(* Logix 5000 project; controller PLC_MCC1300_75F1 vendor 1 type 14 code 166 rev 32.11; software revision 32.04; part 19 of 83 *)
(* tags used below, declared in another part *)
   GP_OB_InitializeMain : GP_OB_Initialize;
   M302SpeedUp : MAC_SpeedUp;
   M310_M4_DR_B1 : AXIS_CIP_DRIVE;
   M310_M5_DR_B2 : AXIS_CIP_DRIVE;
   M310B : MAC_Conveyor;
   M310B_Data : UDT_Convoy_SL;
   M310B_M1_DR_IN_MAR : MOTION_INSTRUCTION;
   M310B_M1_DR_IN_MAS : MOTION_INSTRUCTION;
   M310B_M1_DR_OUT_MAJ : MOTION_INSTRUCTION;
   M310B_M1_DR_OUT_MAS : MOTION_INSTRUCTION;
   M310B_M2_DR_IN_MAJ : MOTION_INSTRUCTION;
   M310B_M2_DR_IN_MAR : MOTION_INSTRUCTION;
   M310B_M2_DR_IN_MAS : MOTION_INSTRUCTION;
   M310B_M2_DR_IN_MRP : MOTION_INSTRUCTION;
   M310B_M2_DR_MAFR : MOTION_INSTRUCTION;
   M310B_M2_DR_MDR : MOTION_INSTRUCTION;
   M310B_M2_DR_MSF : MOTION_INSTRUCTION;
   M310B_M2_DR_MSO : MOTION_INSTRUCTION;
   M310B_M2_DR_OUT_MAJ : MOTION_INSTRUCTION;
   M310B_M2_DR_OUT_MAM : MOTION_INSTRUCTION;
   M310B_M2_DR_OUT_MAR : MOTION_INSTRUCTION;
   M310B_M2_DR_OUT_MAS : MOTION_INSTRUCTION;
   M310B_M2_DR_OUT_MCD : MOTION_INSTRUCTION;
   M310B_M2_DR_OUT_MRP : MOTION_INSTRUCTION;
   M310B_SpaceConv_Utilities : SpaceConv_Utilities;
   M310B_xOS_PosReq : BOOL;
   TMP_d : DINT;
   TMP_dDirection : DINT;
   TMP_r : REAL;
   TMP_rAcc : REAL;
   TMP_rDec : REAL;
   TMP_rSpeed : REAL;
   TMP_rTarget_M2 : REAL;
   TMP_xPositioning : BOOL;
   TMP_xPositioning_M2 : BOOL;
   TMP_xReverse : BOOL;
   TMP_xReverse_M1 : BOOL;
   TMP_xReverse_M2 : BOOL;
   TMP_xRun : BOOL;
   TMP_xRun_M1 : BOOL;
   TMP_xRun_M2 : BOOL;
   xAlwaysOFF : BOOL;
   xDebugOFF : BOOL;
   Z300_Conveyor : UDT_StandConv[29];
   Z300_Conveyor_Conf : UDT_Conveyor_Config[29];
   Z300_Conveyor_HMW : MAC_Conveyor_ZC_HMW[29];
   Z300_Conveyor_IN_MOTION : MAC_Conveyor_ZC_IN_MOTION[29];
   Z301_HMR : MAC_Zone_ML_HMR;
   Z401 : MAC_Zone;
(* CommandLogic, continued *)

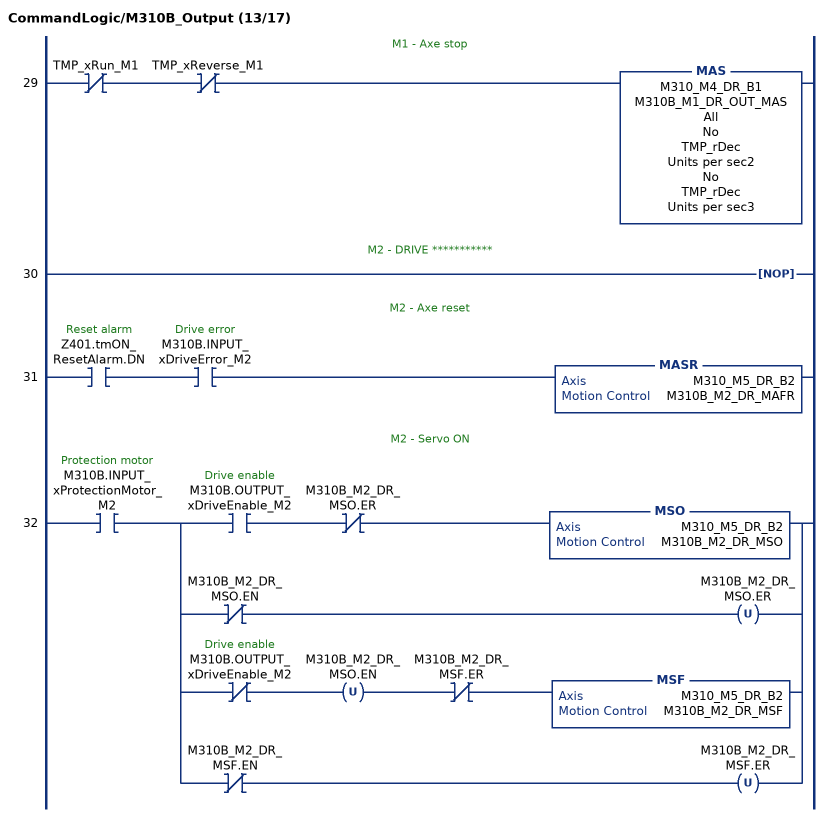
   [picture p150: CommandLogic/M310B_Output rungs 29-32]
   // M1 - Axe stop
   29: XIO(TMP_xRun_M1)XIO(TMP_xReverse_M1)MAS(M310_M4_DR_B1,M310B_M1_DR_OUT_MAS,All,No,TMP_rDec,Units per sec2,No,TMP_rDec,Units per sec3);
   // M2 - DRIVE ***********
   30: NOP();
   // M2 - Axe reset
   31: XIC(Z401.tmON_ResetAlarm.DN)XIC(M310B.INPUT_xDriveError_M2)MASR(M310_M5_DR_B2,M310B_M2_DR_MAFR);
   // M2 - Servo ON
   32: XIC(M310B.INPUT_xProtectionMotor_M2)[XIC(M310B.OUTPUT_xDriveEnable_M2) XIO(M310B_M2_DR_MSO.ER) MSO(M310_M5_DR_B2,M310B_M2_DR_MSO) ,XIO(M310B_M2_DR_MSO.EN) OTU(M310B_M2_DR_MSO.ER) ,XIO(M310B.OUTPUT_xDriveEnable_M2) OTU(M310B_M2_DR_MSO.EN) XIO(M310B_M2_DR_MSF.ER) MSF(M310_M5_DR_B2,M310B_M2_DR_MSF) ,XIO(M310B_M2_DR_MSF.EN) OTU(M310B_M2_DR_MSF.ER) ];
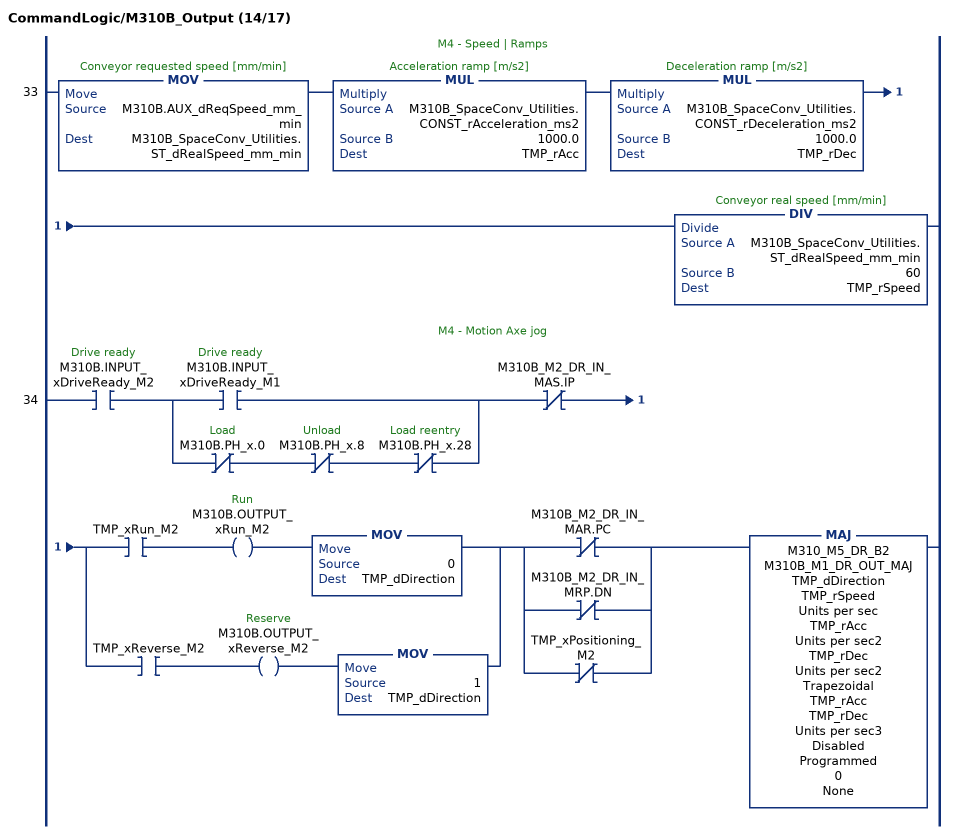
   // M4 - Speed | Ramps
   33: MOV(M310B.AUX_dReqSpeed_mm_min,M310B_SpaceConv_Utilities.ST_dRealSpeed_mm_min)MUL(M310B_SpaceConv_Utilities.CONST_rAcceleration_ms2,1000.0,TMP_rAcc)MUL(M310B_SpaceConv_Utilities.CONST_rDeceleration_ms2,1000.0,TMP_rDec)DIV(M310B_SpaceConv_Utilities.ST_dRealSpeed_mm_min,60,TMP_rSpeed);
   // M4 - Motion Axe jog
   34: XIC(M310B.INPUT_xDriveReady_M2)[XIC(M310B.INPUT_xDriveReady_M1) ,XIO(M310B.PH_x.0) XIO(M310B.PH_x.8) XIO(M310B.PH_x.28) ]XIO(M310B_M2_DR_IN_MAS.IP)[XIC(TMP_xRun_M2) OTE(M310B.OUTPUT_xRun_M2) MOV(0,TMP_dDirection) ,XIC(TMP_xReverse_M2) OTE(M310B.OUTPUT_xReverse_M2) MOV(1,TMP_dDirection) ][XIO(M310B_M2_DR_IN_MAR.PC) ,XIO(M310B_M2_DR_IN_MRP.DN) ,XIO(TMP_xPositioning_M2) ]MAJ(M310_M5_DR_B2,M310B_M1_DR_OUT_MAJ,TMP_dDirection,TMP_rSpeed,Units per sec,TMP_rAcc,Units per sec2,TMP_rDec,Units per sec2,Trapezoidal,TMP_rAcc,TMP_rDec,Units per sec3,Disabled,Programmed,0,None);
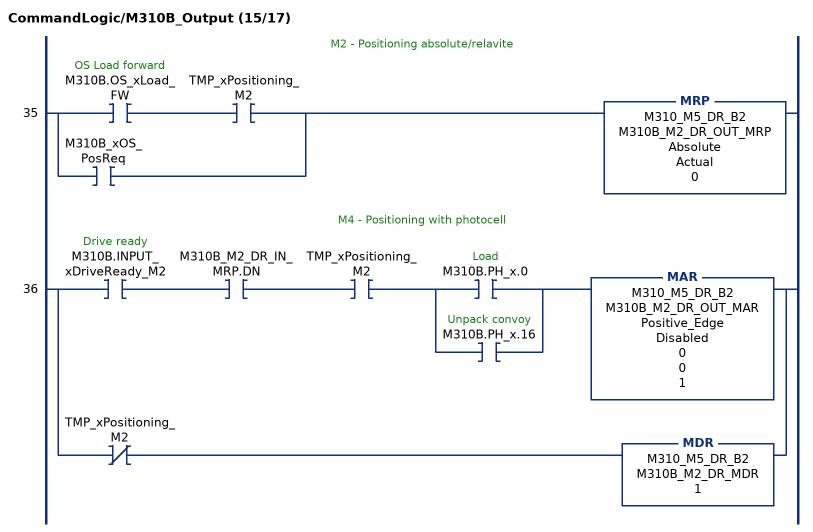
   // M2 - Positioning absolute/relavite
   35: [XIC(M310B.OS_xLoad_FW) XIC(TMP_xPositioning_M2) ,XIC(M310B_xOS_PosReq) ]MRP(M310_M5_DR_B2,M310B_M2_DR_OUT_MRP,Absolute,Actual,0);
   // M4 - Positioning with photocell
   36: [XIC(M310B.INPUT_xDriveReady_M2) XIC(M310B_M2_DR_IN_MRP.DN) XIC(TMP_xPositioning_M2) [XIC(M310B.PH_x.0) ,XIC(M310B.PH_x.16) ] MAR(M310_M5_DR_B2,M310B_M2_DR_OUT_MAR,Positive_Edge,Disabled,0,0,1) ,XIO(TMP_xPositioning_M2) MDR(M310_M5_DR_B2,M310B_M2_DR_MDR,1) ];
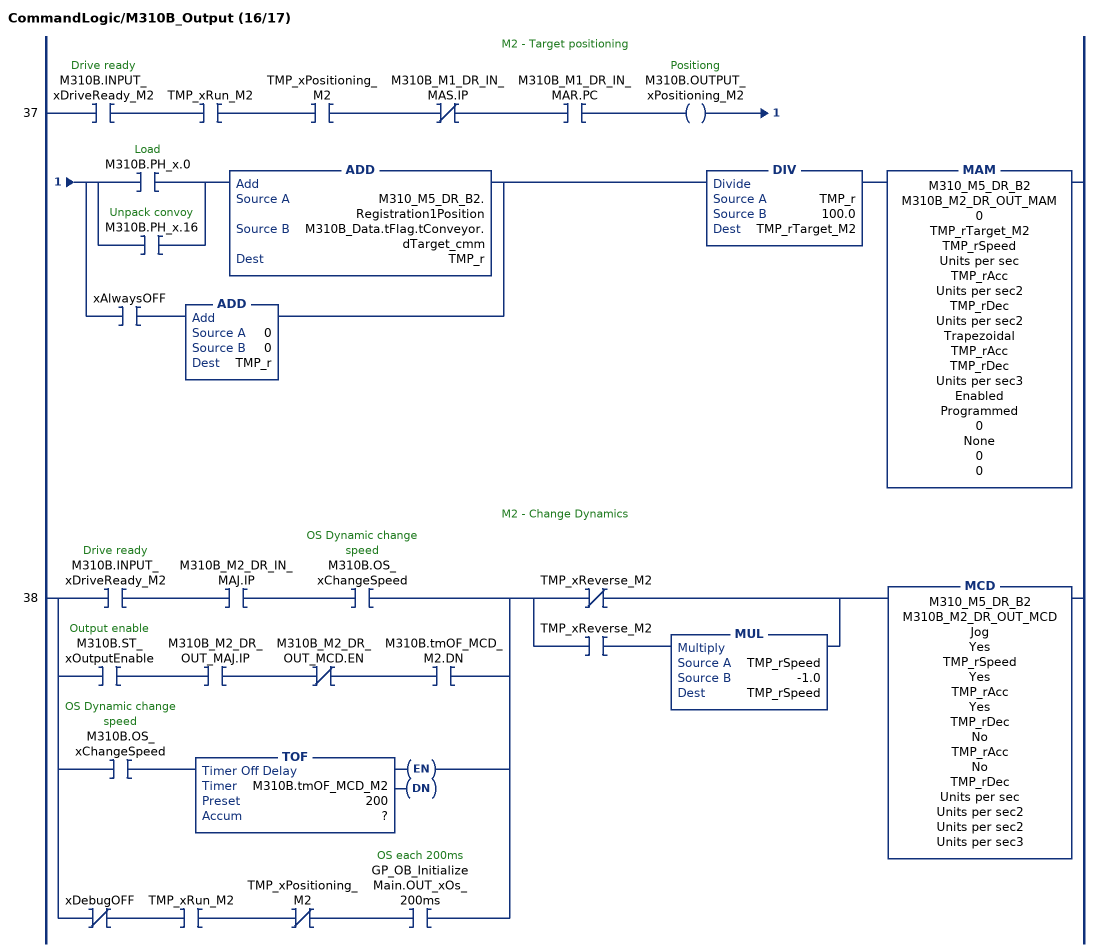
   // M2 - Target positioning
   37: XIC(M310B.INPUT_xDriveReady_M2)XIC(TMP_xRun_M2)XIC(TMP_xPositioning_M2)XIO(M310B_M1_DR_IN_MAS.IP)XIC(M310B_M1_DR_IN_MAR.PC)OTE(M310B.OUTPUT_xPositioning_M2)[[XIC(M310B.PH_x.0) ,XIC(M310B.PH_x.16) ] ADD(M310_M5_DR_B2.Registration1Position,M310B_Data.tFlag.tConveyor.dTarget_cmm,TMP_r) ,XIC(xAlwaysOFF) ADD(0,0,TMP_r) ]DIV(TMP_r,100.0,TMP_rTarget_M2)MAM(M310_M5_DR_B2,M310B_M2_DR_OUT_MAM,0,TMP_rTarget_M2,TMP_rSpeed,Units per sec,TMP_rAcc,Units per sec2,TMP_rDec,Units per sec2,Trapezoidal,TMP_rAcc,TMP_rDec,Units per sec3,Enabled,Programmed,0,None,0,0);
   // M2 - Change Dynamics
   38: [XIC(M310B.INPUT_xDriveReady_M2) XIC(M310B_M2_DR_IN_MAJ.IP) XIC(M310B.OS_xChangeSpeed) ,XIC(M310B.ST_xOutputEnable) XIC(M310B_M2_DR_OUT_MAJ.IP) XIO(M310B_M2_DR_OUT_MCD.EN) XIC(M310B.tmOF_MCD_M2.DN) ,XIC(M310B.OS_xChangeSpeed) TOF(M310B.tmOF_MCD_M2,?,?) ,XIO(xDebugOFF) XIC(TMP_xRun_M2) XIO(TMP_xPositioning_M2) XIC(GP_OB_InitializeMain.OUT_xOs_200ms) ][XIO(TMP_xReverse_M2) ,XIC(TMP_xReverse_M2) MUL(TMP_rSpeed,-1.0,TMP_rSpeed) ]MCD(M310_M5_DR_B2,M310B_M2_DR_OUT_MCD,Jog,Yes,TMP_rSpeed,Yes,TMP_rAcc,Yes,TMP_rDec,No,TMP_rAcc,No,TMP_rDec,Units per sec,Units per sec2,Units per sec2,Units per sec3);
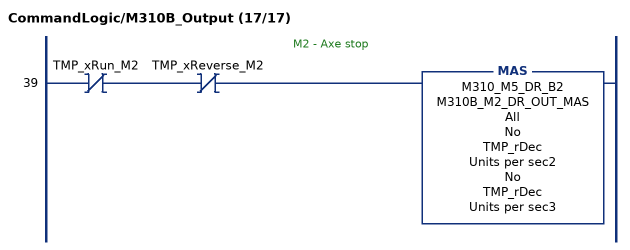
   // M2 - Axe stop
   39: XIO(TMP_xRun_M2)XIO(TMP_xReverse_M2)MAS(M310_M5_DR_B2,M310B_M2_DR_OUT_MAS,All,No,TMP_rDec,Units per sec2,No,TMP_rDec,Units per sec3);
END_ROUTINE

ROUTINE M310M1_Conveyor_Output   (* ladder *)
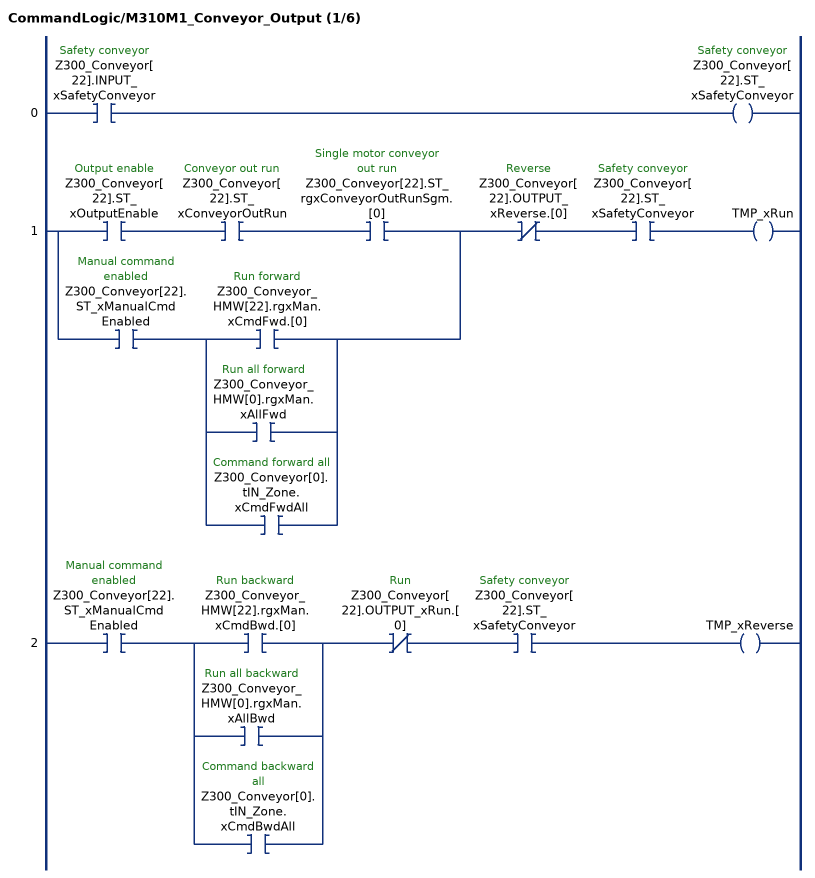
   0: XIC(Z300_Conveyor[22].INPUT_xSafetyConveyor)OTE(Z300_Conveyor[22].ST_xSafetyConveyor);
   1: [XIC(Z300_Conveyor[22].ST_xOutputEnable) XIC(Z300_Conveyor[22].ST_xConveyorOutRun) XIC(Z300_Conveyor[22].ST_rgxConveyorOutRunSgm.[0]) ,XIC(Z300_Conveyor[22].ST_xManualCmdEnabled) [XIC(Z300_Conveyor_HMW[22].rgxMan.xCmdFwd.[0]) ,XIC(Z300_Conveyor_HMW[0].rgxMan.xAllFwd) ,XIC(Z300_Conveyor[0].tIN_Zone.xCmdFwdAll) ] ]XIO(Z300_Conveyor[22].OUTPUT_xReverse.[0])XIC(Z300_Conveyor[22].ST_xSafetyConveyor)OTE(TMP_xRun);
   2: XIC(Z300_Conveyor[22].ST_xManualCmdEnabled)[XIC(Z300_Conveyor_HMW[22].rgxMan.xCmdBwd.[0]) ,XIC(Z300_Conveyor_HMW[0].rgxMan.xAllBwd) ,XIC(Z300_Conveyor[0].tIN_Zone.xCmdBwdAll) ]XIO(Z300_Conveyor[22].OUTPUT_xRun.[0])XIC(Z300_Conveyor[22].ST_xSafetyConveyor)OTE(TMP_xReverse);
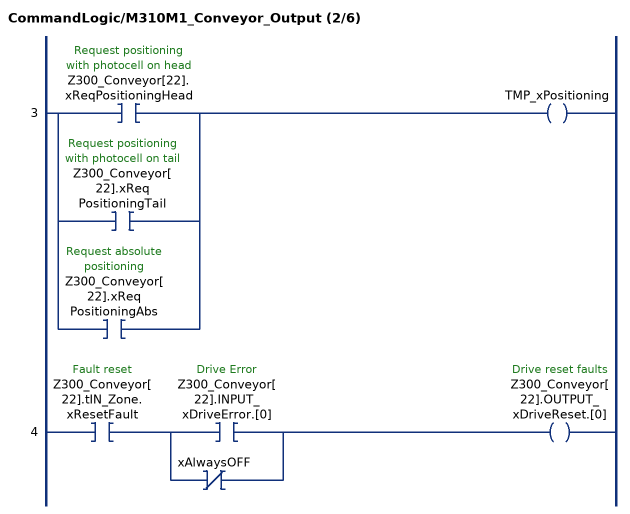
   3: [XIC(Z300_Conveyor[22].xReqPositioningHead) ,XIC(Z300_Conveyor[22].xReqPositioningTail) ,XIC(Z300_Conveyor[22].xReqPositioningAbs) ]OTE(TMP_xPositioning);
   4: XIC(Z300_Conveyor[22].tIN_Zone.xResetFault)[XIC(Z300_Conveyor[22].INPUT_xDriveError.[0]) ,XIO(xAlwaysOFF) ]OTE(Z300_Conveyor[22].OUTPUT_xDriveReset.[0]);
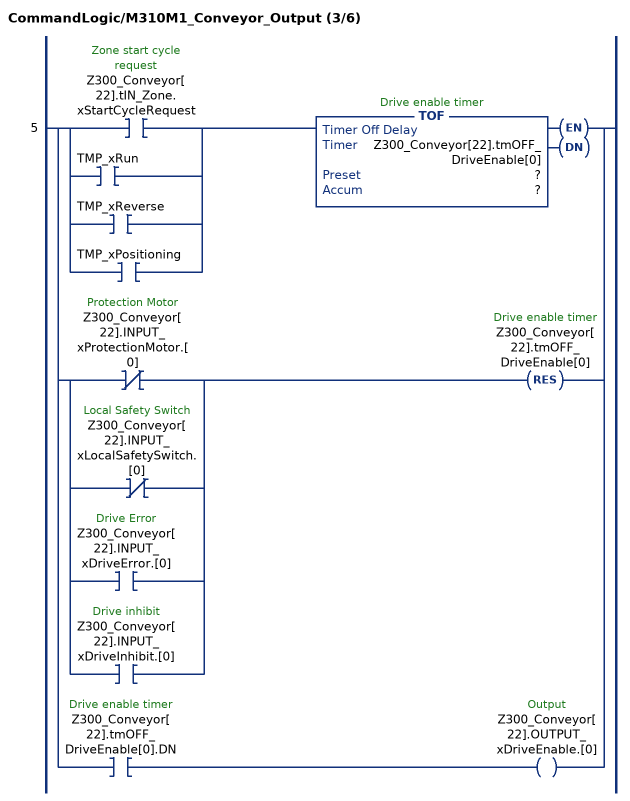
   5: [[XIC(Z300_Conveyor[22].tIN_Zone.xStartCycleRequest) ,XIC(TMP_xRun) ,XIC(TMP_xReverse) ,XIC(TMP_xPositioning) ] TOF(Z300_Conveyor[22].tmOFF_DriveEnable[0],?,?) ,[XIO(Z300_Conveyor[22].INPUT_xProtectionMotor.[0]) ,XIO(Z300_Conveyor[22].INPUT_xLocalSafetySwitch.[0]) ,XIC(Z300_Conveyor[22].INPUT_xDriveError.[0]) ,XIC(Z300_Conveyor[22].INPUT_xDriveInhibit.[0]) ] RES(Z300_Conveyor[22].tmOFF_DriveEnable[0]) ,XIC(Z300_Conveyor[22].tmOFF_DriveEnable[0].DN) OTE(Z300_Conveyor[22].OUTPUT_xDriveEnable.[0]) ];
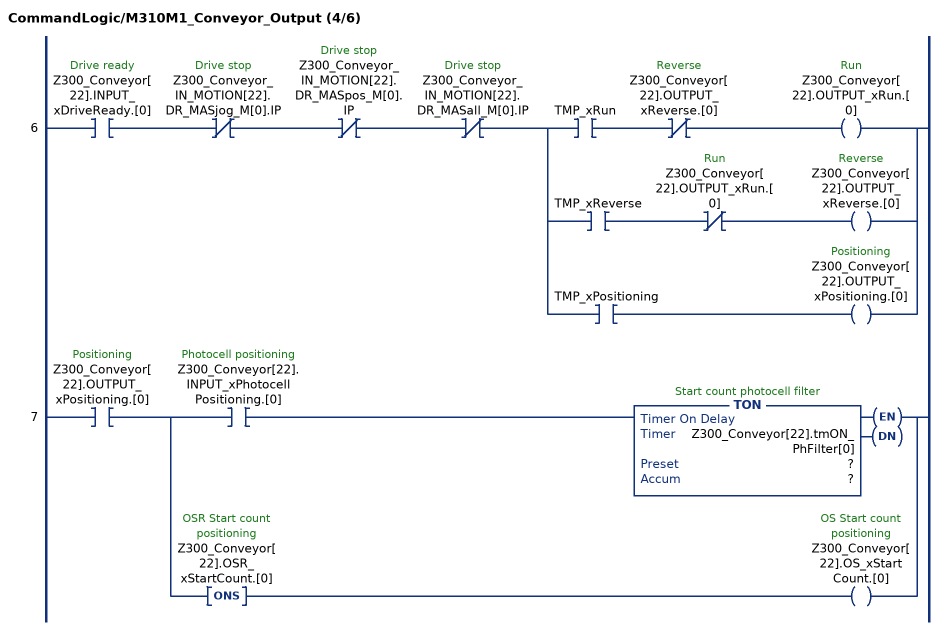
   6: XIC(Z300_Conveyor[22].INPUT_xDriveReady.[0])XIO(Z300_Conveyor_IN_MOTION[22].DR_MASjog_M[0].IP)XIO(Z300_Conveyor_IN_MOTION[22].DR_MASpos_M[0].IP)XIO(Z300_Conveyor_IN_MOTION[22].DR_MASall_M[0].IP)[XIC(TMP_xRun) XIO(Z300_Conveyor[22].OUTPUT_xReverse.[0]) OTE(Z300_Conveyor[22].OUTPUT_xRun.[0]) ,XIC(TMP_xReverse) XIO(Z300_Conveyor[22].OUTPUT_xRun.[0]) OTE(Z300_Conveyor[22].OUTPUT_xReverse.[0]) ,XIC(TMP_xPositioning) OTE(Z300_Conveyor[22].OUTPUT_xPositioning.[0]) ];
   7: XIC(Z300_Conveyor[22].OUTPUT_xPositioning.[0])[XIC(Z300_Conveyor[22].INPUT_xPhotocellPositioning.[0]) TON(Z300_Conveyor[22].tmON_PhFilter[0],?,?) ,ONS(Z300_Conveyor[22].OSR_xStartCount.[0]) OTE(Z300_Conveyor[22].OS_xStartCount.[0]) ];
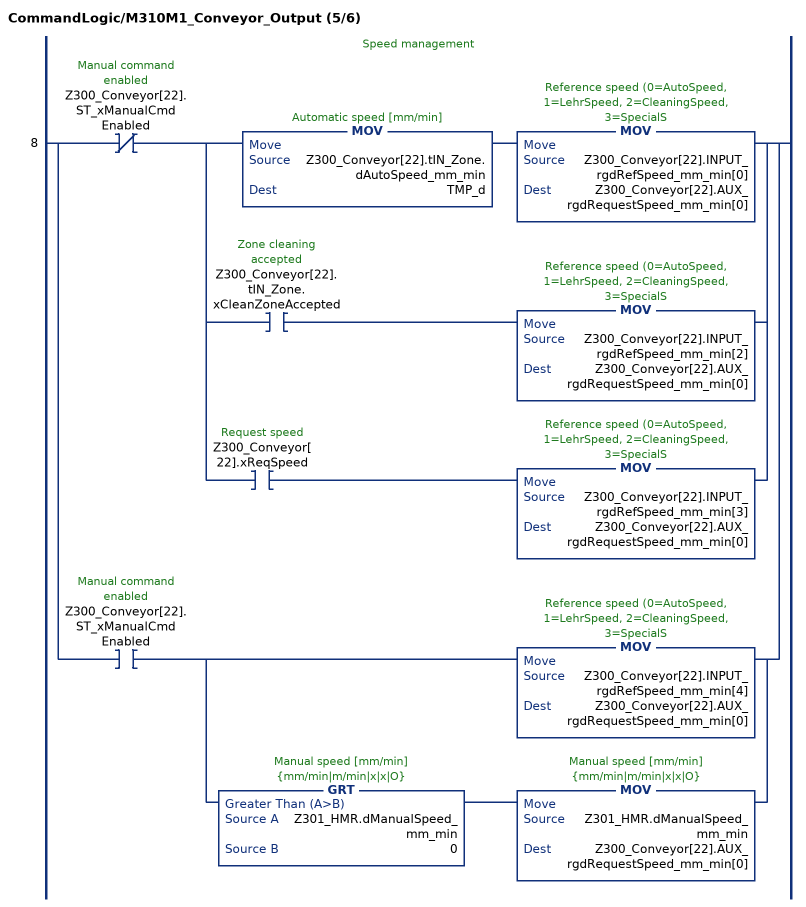
   // Speed management
   8: [XIO(Z300_Conveyor[22].ST_xManualCmdEnabled) [MOV(Z300_Conveyor[22].tIN_Zone.dAutoSpeed_mm_min,TMP_d) MOV(Z300_Conveyor[22].INPUT_rgdRefSpeed_mm_min[0],Z300_Conveyor[22].AUX_rgdRequestSpeed_mm_min[0]) ,XIC(Z300_Conveyor[22].tIN_Zone.xCleanZoneAccepted) MOV(Z300_Conveyor[22].INPUT_rgdRefSpeed_mm_min[2],Z300_Conveyor[22].AUX_rgdRequestSpeed_mm_min[0]) ,XIC(Z300_Conveyor[22].xReqSpeed) MOV(Z300_Conveyor[22].INPUT_rgdRefSpeed_mm_min[3],Z300_Conveyor[22].AUX_rgdRequestSpeed_mm_min[0]) ] ,XIC(Z300_Conveyor[22].ST_xManualCmdEnabled) [MOV(Z300_Conveyor[22].INPUT_rgdRefSpeed_mm_min[4],Z300_Conveyor[22].AUX_rgdRequestSpeed_mm_min[0]) ,GRT(Z301_HMR.dManualSpeed_mm_min,0) MOV(Z301_HMR.dManualSpeed_mm_min,Z300_Conveyor[22].AUX_rgdRequestSpeed_mm_min[0]) ] ];
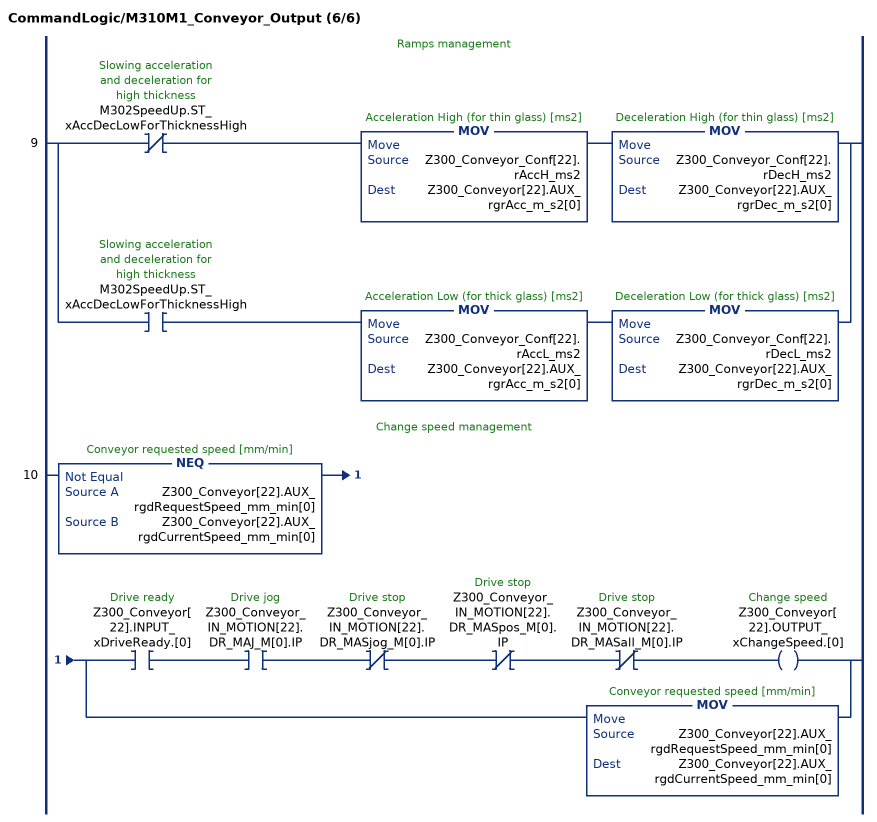
   // Ramps management
   9: [XIO(M302SpeedUp.ST_xAccDecLowForThicknessHigh) MOV(Z300_Conveyor_Conf[22].rAccH_ms2,Z300_Conveyor[22].AUX_rgrAcc_m_s2[0]) MOV(Z300_Conveyor_Conf[22].rDecH_ms2,Z300_Conveyor[22].AUX_rgrDec_m_s2[0]) ,XIC(M302SpeedUp.ST_xAccDecLowForThicknessHigh) MOV(Z300_Conveyor_Conf[22].rAccL_ms2,Z300_Conveyor[22].AUX_rgrAcc_m_s2[0]) MOV(Z300_Conveyor_Conf[22].rDecL_ms2,Z300_Conveyor[22].AUX_rgrDec_m_s2[0]) ];
   // Change speed management
   10: NEQ(Z300_Conveyor[22].AUX_rgdRequestSpeed_mm_min[0],Z300_Conveyor[22].AUX_rgdCurrentSpeed_mm_min[0])[XIC(Z300_Conveyor[22].INPUT_xDriveReady.[0]) XIC(Z300_Conveyor_IN_MOTION[22].DR_MAJ_M[0].IP) XIO(Z300_Conveyor_IN_MOTION[22].DR_MASjog_M[0].IP) XIO(Z300_Conveyor_IN_MOTION[22].DR_MASpos_M[0].IP) XIO(Z300_Conveyor_IN_MOTION[22].DR_MASall_M[0].IP) OTE(Z300_Conveyor[22].OUTPUT_xChangeSpeed.[0]) ,MOV(Z300_Conveyor[22].AUX_rgdRequestSpeed_mm_min[0],Z300_Conveyor[22].AUX_rgdCurrentSpeed_mm_min[0]) ];